REGION Network 34: Send preset command
   RUNG wire#powerrail
      Contact( #STC_tPH.x8 )
      wire#w1
      Contact( #STC_tMngSysReg.tST.xDone )
      wire#w2
      I_Contact( #STC_tMngSysReg.tST.xBusy )
      wire#w3
      I_Contact( #STC_tMngSysReg.tST.xError )
      S_Coil( #STC_tPH.x10 )
   END_RUNG
   RUNG wire#w1
      Contact( #STC_tMngSysReg.tST.xError )
   END_RUNG wire#w2
   RUNG wire#w3
      R_Coil( #STC_tPH.x8 )
   END_RUNG
   // the same network as SCL:
   #_w1 := #STC_tPH.x8 AND (#STC_tMngSysReg.tST.xDone OR #STC_tMngSysReg.tST.xError) AND NOT #STC_tMngSysReg.tST.xBusy;
   IF #_w1 AND NOT #STC_tMngSysReg.tST.xError THEN #STC_tPH.x10 := TRUE; END_IF;
   IF #_w1 THEN #STC_tPH.x8 := FALSE; END_IF;
END_REGION

REGION Network 35 (STL): Error during send ecoder value
         A     #STC_tMngSysReg.tST.xError;
         L     30;
         JC    Err;
END_REGION

REGION Network 36 (STL): Send preset command
         A     #STC_tPH.x10;
         JCN   PrE1;
         =     #STC_tMngSysReg.tST.xWrite_Request;

         L     #STC_tSYS_DATA.iPosPZD_MM;
         +     20;
         SLW   8;
         L     W#16#2;
         OW;
         T     #STC_tMngSysReg.tDATA.wRequest_refere_RequestID;
         L     #STC_tSYS_DATA.iPosPZD_MM;
         SLW   8;
         L     W#16#1;
         OW;
         T     #STC_tMngSysReg.tDATA.wAxis_NoOfParameters;
         L     W#16#1001;
         T     #STC_tMngSysReg.tDATA.wAttribute_NoOfElements;
         L     2507;
         T     #STC_tMngSysReg.tDATA.iParameter_number;
         L     W#16#0;
         T     #STC_tMngSysReg.tDATA.wSubindex;
         L     W#16#4201;
         T     #STC_tMngSysReg.tDATA.wFormat_NoOfValue;
         L     #STC_tSYS_DATA.iDiagAddress;
         T     #STC_tMngSysReg.tST.ID;
         L     47;
         T     #STC_tMngSysReg.tST.dINDEX;
         L     14;
         T     #STC_tMngSysReg.tST.uiLEN;

         L     DINT#2;
         SLD   16;
         T     #STC_tMngSysReg.tDATA.dwRegisterValue;

         CALL  #STC_tWriteRecord
         ( REQ    := #STC_tMngSysReg.tST.xWrite_Request,
           ID     := #STC_tMngSysReg.tST.ID,
           INDEX  := #STC_tMngSysReg.tST.dINDEX,
           LEN    := #STC_tMngSysReg.tST.uiLEN,
           DONE   := #STC_tMngSysReg.tST.xDone,
           BUSY   := #STC_tMngSysReg.tST.xBusy,
           ERROR  := #STC_tMngSysReg.tST.xError,
           STATUS := #STC_tMngSysReg.tST.dwSTATUS,
           RECORD := #STC_tMngSysReg.tDATA
         );
   PrE1: NOP   0;
END_REGION

REGION Network 37: Send saving preset command
   RUNG wire#powerrail
      Contact( #STC_tPH.x10 )
      wire#w1
      Contact( #STC_tMngSysReg.tST.xDone )
      wire#w2
      I_Contact( #STC_tMngSysReg.tST.xBusy )
      wire#w3
      I_Contact( #STC_tMngSysReg.tST.xError )
      S_Coil( #STC_tPH.x12 )
   END_RUNG
   RUNG wire#w1
      Contact( #STC_tMngSysReg.tST.xError )
   END_RUNG wire#w2
   RUNG wire#w3
      R_Coil( #STC_tPH.x10 )
   END_RUNG
   // the same network as SCL:
   #_w1 := #STC_tPH.x10 AND (#STC_tMngSysReg.tST.xDone OR #STC_tMngSysReg.tST.xError) AND NOT #STC_tMngSysReg.tST.xBusy;
   IF #_w1 AND NOT #STC_tMngSysReg.tST.xError THEN #STC_tPH.x12 := TRUE; END_IF;
   IF #_w1 THEN #STC_tPH.x10 := FALSE; END_IF;
END_REGION

REGION Network 38 (STL): Error during preset command
         A     #STC_tMngSysReg.tST.xError;
         L     31;
         JC    Err;
END_REGION

REGION Network 39 (STL): Send saving preset command
         A     #STC_tPH.x12;
         JCN   PrE2;
         =     #STC_tMngSysReg.tST.xWrite_Request;

         L     #STC_tSYS_DATA.iPosPZD_MM;
         +     30;
         SLW   8;
         L     W#16#2;
         OW;
         T     #STC_tMngSysReg.tDATA.wRequest_refere_RequestID;
         L     #STC_tSYS_DATA.iPosPZD_CU;
         SLW   8;
         L     W#16#1;
         OW;
         T     #STC_tMngSysReg.tDATA.wAxis_NoOfParameters;
         L     W#16#1001;
         T     #STC_tMngSysReg.tDATA.wAttribute_NoOfElements;
         L     977;
         T     #STC_tMngSysReg.tDATA.iParameter_number;
         L     W#16#0;
         T     #STC_tMngSysReg.tDATA.wSubindex;
         L     W#16#4201;
         T     #STC_tMngSysReg.tDATA.wFormat_NoOfValue;
         L     #STC_tSYS_DATA.iDiagAddress;
         T     #STC_tMngSysReg.tST.ID;
         L     47;
         T     #STC_tMngSysReg.tST.dINDEX;
         L     14;
         T     #STC_tMngSysReg.tST.uiLEN;

         L     DINT#1;
         SLD   16;
         T     #STC_tMngSysReg.tDATA.dwRegisterValue;

         CALL  #STC_tWriteRecord
         ( REQ    := #STC_tMngSysReg.tST.xWrite_Request,
           ID     := #STC_tMngSysReg.tST.ID,
           INDEX  := #STC_tMngSysReg.tST.dINDEX,
           LEN    := #STC_tMngSysReg.tST.uiLEN,
           DONE   := #STC_tMngSysReg.tST.xDone,
           BUSY   := #STC_tMngSysReg.tST.xBusy,
           ERROR  := #STC_tMngSysReg.tST.xError,
           STATUS := #STC_tMngSysReg.tST.dwSTATUS,
           RECORD := #STC_tMngSysReg.tDATA
         );
   PrE2: NOP   0;
END_REGION

REGION Network 40: End preset encoder
   RUNG wire#powerrail
      Contact( #STC_tPH.x12 )
      wire#w1
      Contact( #STC_tMngSysReg.tST.xDone )
      wire#w2
      I_Contact( #STC_tMngSysReg.tST.xBusy )
      wire#w3
      Coil( #STC_tPH.x14 )
   END_RUNG
   RUNG wire#w1
      Contact( #STC_tMngSysReg.tST.xError )
   END_RUNG wire#w2
   RUNG wire#w3
      R_Coil( #STC_tPH.x12 )
   END_RUNG
   // the same network as SCL:
   #STC_tPH.x14 := #STC_tPH.x12 AND (#STC_tMngSysReg.tST.xDone OR #STC_tMngSysReg.tST.xError) AND NOT #STC_tMngSysReg.tST.xBusy;
   IF #STC_tPH.x14 THEN #STC_tPH.x12 := FALSE; END_IF;
END_REGION

REGION Network 41 (STL): Error during saving preset command
         A     #STC_tMngSysReg.tST.xError;
         L     32;
         JC    Err;
END_REGION

REGION Network 42: Preset phases in progress
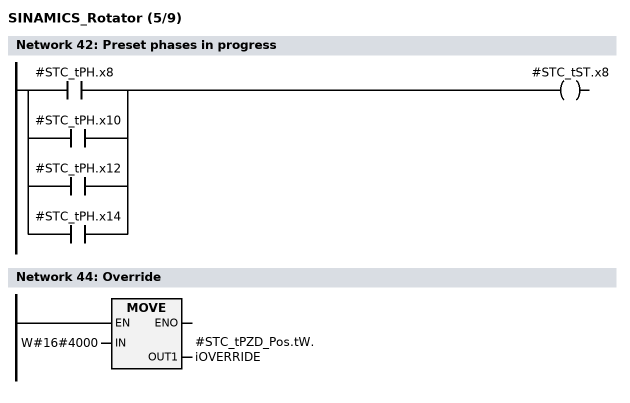
   RUNG wire#powerrail
      Contact( #STC_tPH.x8 )
      wire#w1
      Coil( #STC_tST.x8 )
   END_RUNG
   RUNG wire#powerrail
      Contact( #STC_tPH.x10 )
   END_RUNG wire#w1
   RUNG wire#powerrail
      Contact( #STC_tPH.x12 )
   END_RUNG wire#w1
   RUNG wire#powerrail
      Contact( #STC_tPH.x14 )
   END_RUNG wire#w1
   // the same network as SCL:
   #STC_tST.x8 := #STC_tPH.x8 OR #STC_tPH.x10 OR #STC_tPH.x12 OR #STC_tPH.x14;
END_REGION

REGION Network 43: #####_PARAMETERS_#####
END_REGION

REGION Network 44: Override
   RUNG wire#powerrail
      { S7_GenerateENO := "TRUE" } Move(in := W#16#4000, out1 => #STC_tPZD_Pos.tW.iOVERRIDE)
   END_RUNG
   // the same network as SCL:
   #STC_tPZD_Pos.tW.iOVERRIDE := W#16#4000;
END_REGION

REGION Network 45: Actual position filtered
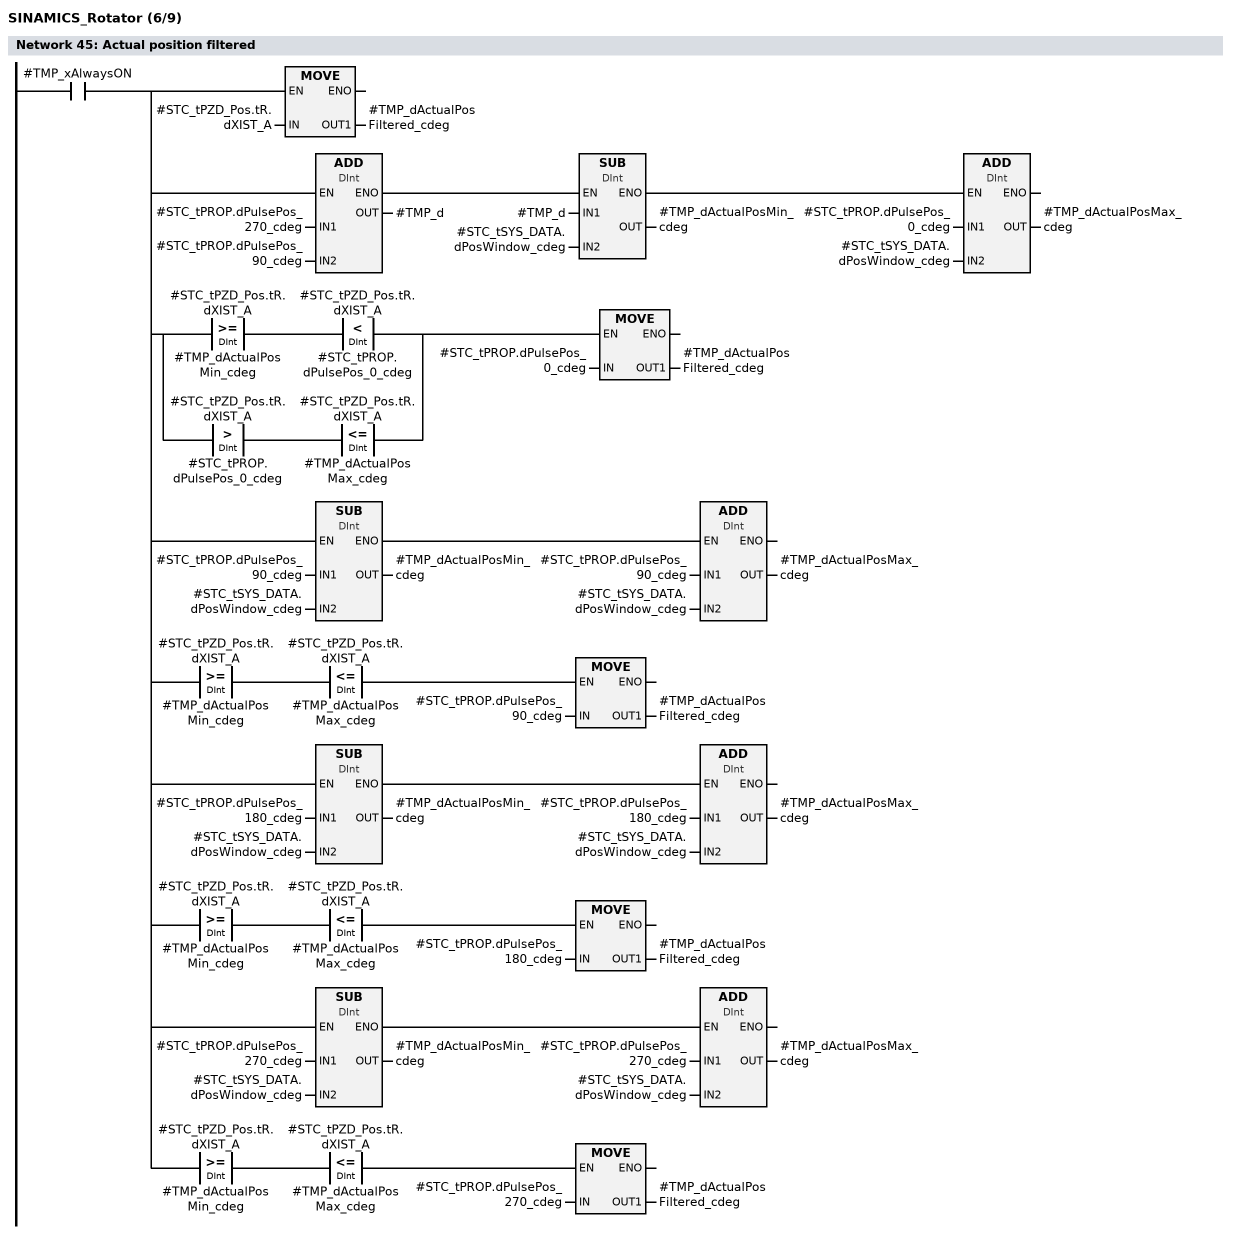
   RUNG wire#powerrail
      Contact( #TMP_xAlwaysON )
      wire#w1
      { S7_GenerateENO := "TRUE" } Move(in := #STC_tPZD_Pos.tR.dXIST_A, out1 => #TMP_dActualPosFiltered_cdeg)
   END_RUNG
   RUNG wire#w1
      { S7_Templates := "SrcType := DInt"; S7_GenerateENO := "TRUE" } Add(in1 := #STC_tPROP.dPulsePos_270_cdeg, in2 := #STC_tPROP.dPulsePos_90_cdeg, out => #TMP_d)
      { S7_Templates := "SrcType := DInt"; S7_GenerateENO := "TRUE" } Sub(in1 := #TMP_d, in2 := #STC_tSYS_DATA.dPosWindow_cdeg, out => #TMP_dActualPosMin_cdeg)
      { S7_Templates := "SrcType := DInt"; S7_GenerateENO := "TRUE" } Add(in1 := #STC_tPROP.dPulsePos_0_cdeg, in2 := #STC_tSYS_DATA.dPosWindow_cdeg, out => #TMP_dActualPosMax_cdeg)
   END_RUNG
   RUNG wire#w1
      { S7_Templates := "SrcType := DInt" } GE_Contact(in1 := #STC_tPZD_Pos.tR.dXIST_A, in2 := #TMP_dActualPosMin_cdeg)
      { S7_Templates := "SrcType := DInt" } LT_Contact(in1 := #STC_tPZD_Pos.tR.dXIST_A, in2 := #STC_tPROP.dPulsePos_0_cdeg)
      wire#w2
      { S7_GenerateENO := "TRUE" } Move(in := #STC_tPROP.dPulsePos_0_cdeg, out1 => #TMP_dActualPosFiltered_cdeg)
   END_RUNG
   RUNG wire#w1
      { S7_Templates := "SrcType := DInt" } GT_Contact(in1 := #STC_tPZD_Pos.tR.dXIST_A, in2 := #STC_tPROP.dPulsePos_0_cdeg)
      { S7_Templates := "SrcType := DInt" } LE_Contact(in1 := #STC_tPZD_Pos.tR.dXIST_A, in2 := #TMP_dActualPosMax_cdeg)
   END_RUNG wire#w2
   RUNG wire#w1
      { S7_Templates := "SrcType := DInt"; S7_GenerateENO := "TRUE" } Sub(in1 := #STC_tPROP.dPulsePos_90_cdeg, in2 := #STC_tSYS_DATA.dPosWindow_cdeg, out => #TMP_dActualPosMin_cdeg)
      { S7_Templates := "SrcType := DInt"; S7_GenerateENO := "TRUE" } Add(in1 := #STC_tPROP.dPulsePos_90_cdeg, in2 := #STC_tSYS_DATA.dPosWindow_cdeg, out => #TMP_dActualPosMax_cdeg)
   END_RUNG
   RUNG wire#w1
      { S7_Templates := "SrcType := DInt" } GE_Contact(in1 := #STC_tPZD_Pos.tR.dXIST_A, in2 := #TMP_dActualPosMin_cdeg)
      { S7_Templates := "SrcType := DInt" } LE_Contact(in1 := #STC_tPZD_Pos.tR.dXIST_A, in2 := #TMP_dActualPosMax_cdeg)
      { S7_GenerateENO := "TRUE" } Move(in := #STC_tPROP.dPulsePos_90_cdeg, out1 => #TMP_dActualPosFiltered_cdeg)
   END_RUNG
   RUNG wire#w1
      { S7_Templates := "SrcType := DInt"; S7_GenerateENO := "TRUE" } Sub(in1 := #STC_tPROP.dPulsePos_180_cdeg, in2 := #STC_tSYS_DATA.dPosWindow_cdeg, out => #TMP_dActualPosMin_cdeg)
      { S7_Templates := "SrcType := DInt"; S7_GenerateENO := "TRUE" } Add(in1 := #STC_tPROP.dPulsePos_180_cdeg, in2 := #STC_tSYS_DATA.dPosWindow_cdeg, out => #TMP_dActualPosMax_cdeg)
   END_RUNG
   RUNG wire#w1
      { S7_Templates := "SrcType := DInt" } GE_Contact(in1 := #STC_tPZD_Pos.tR.dXIST_A, in2 := #TMP_dActualPosMin_cdeg)
      { S7_Templates := "SrcType := DInt" } LE_Contact(in1 := #STC_tPZD_Pos.tR.dXIST_A, in2 := #TMP_dActualPosMax_cdeg)
      { S7_GenerateENO := "TRUE" } Move(in := #STC_tPROP.dPulsePos_180_cdeg, out1 => #TMP_dActualPosFiltered_cdeg)
   END_RUNG
   RUNG wire#w1
      { S7_Templates := "SrcType := DInt"; S7_GenerateENO := "TRUE" } Sub(in1 := #STC_tPROP.dPulsePos_270_cdeg, in2 := #STC_tSYS_DATA.dPosWindow_cdeg, out => #TMP_dActualPosMin_cdeg)
      { S7_Templates := "SrcType := DInt"; S7_GenerateENO := "TRUE" } Add(in1 := #STC_tPROP.dPulsePos_270_cdeg, in2 := #STC_tSYS_DATA.dPosWindow_cdeg, out => #TMP_dActualPosMax_cdeg)
   END_RUNG
   RUNG wire#w1
      { S7_Templates := "SrcType := DInt" } GE_Contact(in1 := #STC_tPZD_Pos.tR.dXIST_A, in2 := #TMP_dActualPosMin_cdeg)
      { S7_Templates := "SrcType := DInt" } LE_Contact(in1 := #STC_tPZD_Pos.tR.dXIST_A, in2 := #TMP_dActualPosMax_cdeg)
      { S7_GenerateENO := "TRUE" } Move(in := #STC_tPROP.dPulsePos_270_cdeg, out1 => #TMP_dActualPosFiltered_cdeg)
   END_RUNG
   // the same network as SCL:
   // ENO of a box is taken as its EN; it also drops when the box reports an error
   IF #TMP_xAlwaysON THEN
       #TMP_dActualPosFiltered_cdeg := #STC_tPZD_Pos.tR.dXIST_A;
       #TMP_d := #STC_tPROP.dPulsePos_270_cdeg + #STC_tPROP.dPulsePos_90_cdeg;
       #TMP_dActualPosMin_cdeg := #TMP_d - #STC_tSYS_DATA.dPosWindow_cdeg;
       #TMP_dActualPosMax_cdeg := #STC_tPROP.dPulsePos_0_cdeg + #STC_tSYS_DATA.dPosWindow_cdeg;
   END_IF;
   IF #TMP_xAlwaysON AND (((#STC_tPZD_Pos.tR.dXIST_A >= #TMP_dActualPosMin_cdeg) AND (#STC_tPZD_Pos.tR.dXIST_A < #STC_tPROP.dPulsePos_0_cdeg)) OR ((#STC_tPZD_Pos.tR.dXIST_A > #STC_tPROP.dPulsePos_0_cdeg) AND (#STC_tPZD_Pos.tR.dXIST_A <= #TMP_dActualPosMax_cdeg))) THEN
       #TMP_dActualPosFiltered_cdeg := #STC_tPROP.dPulsePos_0_cdeg;
   END_IF;
   IF #TMP_xAlwaysON THEN
       #TMP_dActualPosMin_cdeg := #STC_tPROP.dPulsePos_90_cdeg - #STC_tSYS_DATA.dPosWindow_cdeg;
       #TMP_dActualPosMax_cdeg := #STC_tPROP.dPulsePos_90_cdeg + #STC_tSYS_DATA.dPosWindow_cdeg;
   END_IF;
   IF #TMP_xAlwaysON AND (#STC_tPZD_Pos.tR.dXIST_A >= #TMP_dActualPosMin_cdeg) AND (#STC_tPZD_Pos.tR.dXIST_A <= #TMP_dActualPosMax_cdeg) THEN
       #TMP_dActualPosFiltered_cdeg := #STC_tPROP.dPulsePos_90_cdeg;
   END_IF;
   IF #TMP_xAlwaysON THEN
       #TMP_dActualPosMin_cdeg := #STC_tPROP.dPulsePos_180_cdeg - #STC_tSYS_DATA.dPosWindow_cdeg;
       #TMP_dActualPosMax_cdeg := #STC_tPROP.dPulsePos_180_cdeg + #STC_tSYS_DATA.dPosWindow_cdeg;
   END_IF;
   IF #TMP_xAlwaysON AND (#STC_tPZD_Pos.tR.dXIST_A >= #TMP_dActualPosMin_cdeg) AND (#STC_tPZD_Pos.tR.dXIST_A <= #TMP_dActualPosMax_cdeg) THEN
       #TMP_dActualPosFiltered_cdeg := #STC_tPROP.dPulsePos_180_cdeg;
   END_IF;
   IF #TMP_xAlwaysON THEN
       #TMP_dActualPosMin_cdeg := #STC_tPROP.dPulsePos_270_cdeg - #STC_tSYS_DATA.dPosWindow_cdeg;
       #TMP_dActualPosMax_cdeg := #STC_tPROP.dPulsePos_270_cdeg + #STC_tSYS_DATA.dPosWindow_cdeg;
   END_IF;
   IF #TMP_xAlwaysON AND (#STC_tPZD_Pos.tR.dXIST_A >= #TMP_dActualPosMin_cdeg) AND (#STC_tPZD_Pos.tR.dXIST_A <= #TMP_dActualPosMax_cdeg) THEN
       #TMP_dActualPosFiltered_cdeg := #STC_tPROP.dPulsePos_270_cdeg;
   END_IF;
END_REGION

REGION Network 46: Target selection
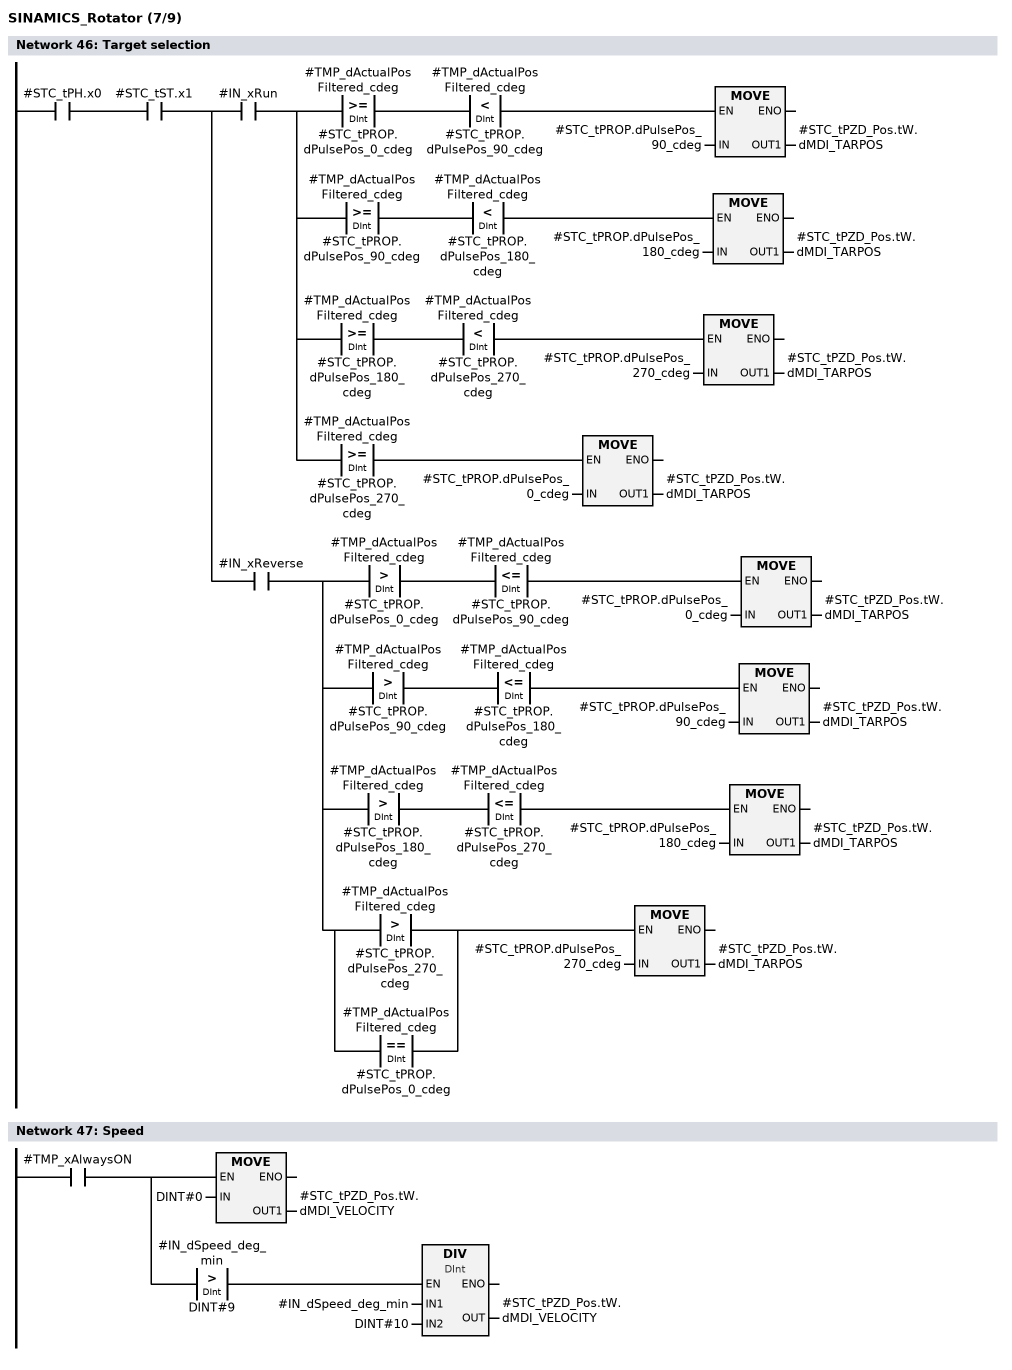
   RUNG wire#powerrail
      Contact( #STC_tPH.x0 )
      Contact( #STC_tST.x1 )
      wire#w1
      Contact( #IN_xRun )
      wire#w2
      { S7_Templates := "SrcType := DInt" } GE_Contact(in1 := #TMP_dActualPosFiltered_cdeg, in2 := #STC_tPROP.dPulsePos_0_cdeg)
      { S7_Templates := "SrcType := DInt" } LT_Contact(in1 := #TMP_dActualPosFiltered_cdeg, in2 := #STC_tPROP.dPulsePos_90_cdeg)
      { S7_GenerateENO := "TRUE" } Move(in := #STC_tPROP.dPulsePos_90_cdeg, out1 => #STC_tPZD_Pos.tW.dMDI_TARPOS)
   END_RUNG
   RUNG wire#w2
      { S7_Templates := "SrcType := DInt" } GE_Contact(in1 := #TMP_dActualPosFiltered_cdeg, in2 := #STC_tPROP.dPulsePos_90_cdeg)
      { S7_Templates := "SrcType := DInt" } LT_Contact(in1 := #TMP_dActualPosFiltered_cdeg, in2 := #STC_tPROP.dPulsePos_180_cdeg)
      { S7_GenerateENO := "TRUE" } Move(in := #STC_tPROP.dPulsePos_180_cdeg, out1 => #STC_tPZD_Pos.tW.dMDI_TARPOS)
   END_RUNG
   RUNG wire#w2
      { S7_Templates := "SrcType := DInt" } GE_Contact(in1 := #TMP_dActualPosFiltered_cdeg, in2 := #STC_tPROP.dPulsePos_180_cdeg)
      { S7_Templates := "SrcType := DInt" } LT_Contact(in1 := #TMP_dActualPosFiltered_cdeg, in2 := #STC_tPROP.dPulsePos_270_cdeg)
      { S7_GenerateENO := "TRUE" } Move(in := #STC_tPROP.dPulsePos_270_cdeg, out1 => #STC_tPZD_Pos.tW.dMDI_TARPOS)
   END_RUNG
   RUNG wire#w2
      { S7_Templates := "SrcType := DInt" } GE_Contact(in1 := #TMP_dActualPosFiltered_cdeg, in2 := #STC_tPROP.dPulsePos_270_cdeg)
      { S7_GenerateENO := "TRUE" } Move(in := #STC_tPROP.dPulsePos_0_cdeg, out1 => #STC_tPZD_Pos.tW.dMDI_TARPOS)
   END_RUNG
   RUNG wire#w1
      Contact( #IN_xReverse )
      wire#w3
      { S7_Templates := "SrcType := DInt" } GT_Contact(in1 := #TMP_dActualPosFiltered_cdeg, in2 := #STC_tPROP.dPulsePos_0_cdeg)
      { S7_Templates := "SrcType := DInt" } LE_Contact(in1 := #TMP_dActualPosFiltered_cdeg, in2 := #STC_tPROP.dPulsePos_90_cdeg)
      { S7_GenerateENO := "TRUE" } Move(in := #STC_tPROP.dPulsePos_0_cdeg, out1 => #STC_tPZD_Pos.tW.dMDI_TARPOS)
   END_RUNG
   RUNG wire#w3
      { S7_Templates := "SrcType := DInt" } GT_Contact(in1 := #TMP_dActualPosFiltered_cdeg, in2 := #STC_tPROP.dPulsePos_90_cdeg)
      { S7_Templates := "SrcType := DInt" } LE_Contact(in1 := #TMP_dActualPosFiltered_cdeg, in2 := #STC_tPROP.dPulsePos_180_cdeg)
      { S7_GenerateENO := "TRUE" } Move(in := #STC_tPROP.dPulsePos_90_cdeg, out1 => #STC_tPZD_Pos.tW.dMDI_TARPOS)
   END_RUNG
   RUNG wire#w3
      { S7_Templates := "SrcType := DInt" } GT_Contact(in1 := #TMP_dActualPosFiltered_cdeg, in2 := #STC_tPROP.dPulsePos_180_cdeg)
      { S7_Templates := "SrcType := DInt" } LE_Contact(in1 := #TMP_dActualPosFiltered_cdeg, in2 := #STC_tPROP.dPulsePos_270_cdeg)
      { S7_GenerateENO := "TRUE" } Move(in := #STC_tPROP.dPulsePos_180_cdeg, out1 => #STC_tPZD_Pos.tW.dMDI_TARPOS)
   END_RUNG
   RUNG wire#w3
      { S7_Templates := "SrcType := DInt" } GT_Contact(in1 := #TMP_dActualPosFiltered_cdeg, in2 := #STC_tPROP.dPulsePos_270_cdeg)
      wire#w4
      { S7_GenerateENO := "TRUE" } Move(in := #STC_tPROP.dPulsePos_270_cdeg, out1 => #STC_tPZD_Pos.tW.dMDI_TARPOS)
   END_RUNG
   RUNG wire#w3
      { S7_Templates := "SrcType := DInt" } EQ_Contact(in1 := #TMP_dActualPosFiltered_cdeg, in2 := #STC_tPROP.dPulsePos_0_cdeg)
   END_RUNG wire#w4
   // the same network as SCL:
   #_w1 := #STC_tPH.x0 AND #STC_tST.x1;
   #_w2 := #_w1 AND #IN_xRun;
   IF #_w2 AND (#TMP_dActualPosFiltered_cdeg >= #STC_tPROP.dPulsePos_0_cdeg) AND (#TMP_dActualPosFiltered_cdeg < #STC_tPROP.dPulsePos_90_cdeg) THEN
       #STC_tPZD_Pos.tW.dMDI_TARPOS := #STC_tPROP.dPulsePos_90_cdeg;
   END_IF;
   IF #_w2 AND (#TMP_dActualPosFiltered_cdeg >= #STC_tPROP.dPulsePos_90_cdeg) AND (#TMP_dActualPosFiltered_cdeg < #STC_tPROP.dPulsePos_180_cdeg) THEN
       #STC_tPZD_Pos.tW.dMDI_TARPOS := #STC_tPROP.dPulsePos_180_cdeg;
   END_IF;
   IF #_w2 AND (#TMP_dActualPosFiltered_cdeg >= #STC_tPROP.dPulsePos_180_cdeg) AND (#TMP_dActualPosFiltered_cdeg < #STC_tPROP.dPulsePos_270_cdeg) THEN
       #STC_tPZD_Pos.tW.dMDI_TARPOS := #STC_tPROP.dPulsePos_270_cdeg;
   END_IF;
   IF #_w2 AND (#TMP_dActualPosFiltered_cdeg >= #STC_tPROP.dPulsePos_270_cdeg) THEN
       #STC_tPZD_Pos.tW.dMDI_TARPOS := #STC_tPROP.dPulsePos_0_cdeg;
   END_IF;
   #_w3 := #_w1 AND #IN_xReverse;
   IF #_w3 AND (#TMP_dActualPosFiltered_cdeg > #STC_tPROP.dPulsePos_0_cdeg) AND (#TMP_dActualPosFiltered_cdeg <= #STC_tPROP.dPulsePos_90_cdeg) THEN
       #STC_tPZD_Pos.tW.dMDI_TARPOS := #STC_tPROP.dPulsePos_0_cdeg;
   END_IF;
   IF #_w3 AND (#TMP_dActualPosFiltered_cdeg > #STC_tPROP.dPulsePos_90_cdeg) AND (#TMP_dActualPosFiltered_cdeg <= #STC_tPROP.dPulsePos_180_cdeg) THEN
       #STC_tPZD_Pos.tW.dMDI_TARPOS := #STC_tPROP.dPulsePos_90_cdeg;
   END_IF;
   IF #_w3 AND (#TMP_dActualPosFiltered_cdeg > #STC_tPROP.dPulsePos_180_cdeg) AND (#TMP_dActualPosFiltered_cdeg <= #STC_tPROP.dPulsePos_270_cdeg) THEN
       #STC_tPZD_Pos.tW.dMDI_TARPOS := #STC_tPROP.dPulsePos_180_cdeg;
   END_IF;
   IF #_w3 AND ((#TMP_dActualPosFiltered_cdeg > #STC_tPROP.dPulsePos_270_cdeg) OR (#TMP_dActualPosFiltered_cdeg = #STC_tPROP.dPulsePos_0_cdeg)) THEN
       #STC_tPZD_Pos.tW.dMDI_TARPOS := #STC_tPROP.dPulsePos_270_cdeg;
   END_IF;
END_REGION

REGION Network 47: Speed
   RUNG wire#powerrail
      Contact( #TMP_xAlwaysON )
      wire#w1
      { S7_GenerateENO := "TRUE" } Move(in := DINT#0, out1 => #STC_tPZD_Pos.tW.dMDI_VELOCITY)
   END_RUNG
   RUNG wire#w1
      { S7_Templates := "SrcType := DInt" } GT_Contact(in1 := #IN_dSpeed_deg_min, in2 := DINT#9)
      { S7_Templates := "SrcType := DInt"; S7_GenerateENO := "TRUE" } Div(in1 := #IN_dSpeed_deg_min, in2 := DINT#10, out => #STC_tPZD_Pos.tW.dMDI_VELOCITY)
   END_RUNG
   // the same network as SCL:
   IF #TMP_xAlwaysON THEN #STC_tPZD_Pos.tW.dMDI_VELOCITY := DINT#0; END_IF;
   IF #TMP_xAlwaysON AND (#IN_dSpeed_deg_min > DINT#9) THEN
       #STC_tPZD_Pos.tW.dMDI_VELOCITY := #IN_dSpeed_deg_min / DINT#10;
   END_IF;
END_REGION

REGION Network 48: Acceleration
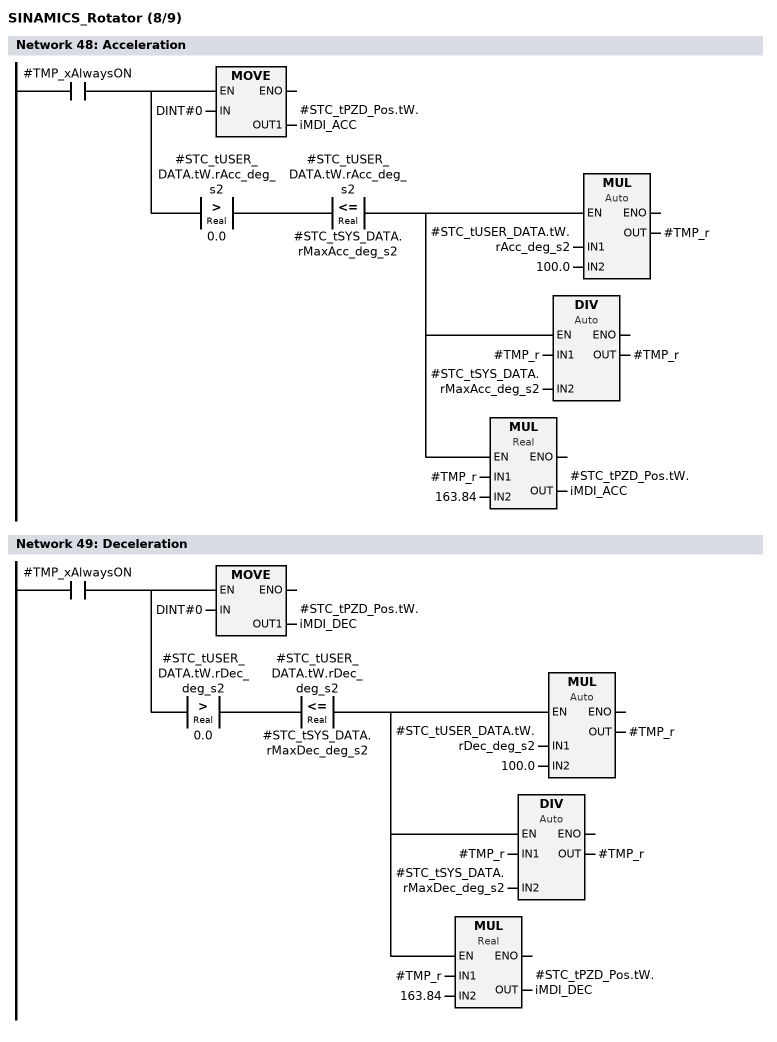
   RUNG wire#powerrail
      Contact( #TMP_xAlwaysON )
      wire#w1
      Move(in := DINT#0, out1 => #STC_tPZD_Pos.tW.iMDI_ACC)
   END_RUNG
   RUNG wire#w1
      { S7_Templates := "SrcType := Real" } GT_Contact(in1 := #STC_tUSER_DATA.tW.rAcc_deg_s2, in2 := 0.0)
      { S7_Templates := "SrcType := Real" } LE_Contact(in1 := #STC_tUSER_DATA.tW.rAcc_deg_s2, in2 := #STC_tSYS_DATA.rMaxAcc_deg_s2)
      wire#w2
      Mul(in1 := #STC_tUSER_DATA.tW.rAcc_deg_s2, in2 := 100.0, out => #TMP_r)
   END_RUNG
   RUNG wire#w2
      Div(in1 := #TMP_r, in2 := #STC_tSYS_DATA.rMaxAcc_deg_s2, out => #TMP_r)
   END_RUNG
   RUNG wire#w2
      { S7_Templates := "SrcType := Real" } Mul(in1 := #TMP_r, in2 := 163.84, out => #STC_tPZD_Pos.tW.iMDI_ACC)
   END_RUNG
   // the same network as SCL:
   IF #TMP_xAlwaysON THEN #STC_tPZD_Pos.tW.iMDI_ACC := DINT#0; END_IF;
   IF #TMP_xAlwaysON AND (#STC_tUSER_DATA.tW.rAcc_deg_s2 > 0.0) AND (#STC_tUSER_DATA.tW.rAcc_deg_s2 <= #STC_tSYS_DATA.rMaxAcc_deg_s2) THEN
       #TMP_r := #STC_tUSER_DATA.tW.rAcc_deg_s2 * 100.0;
       #TMP_r := #TMP_r / #STC_tSYS_DATA.rMaxAcc_deg_s2;
       #STC_tPZD_Pos.tW.iMDI_ACC := #TMP_r * 163.84;
   END_IF;
END_REGION

REGION Network 49: Deceleration
   RUNG wire#powerrail
      Contact( #TMP_xAlwaysON )
      wire#w1
      Move(in := DINT#0, out1 => #STC_tPZD_Pos.tW.iMDI_DEC)
   END_RUNG
   RUNG wire#w1
      { S7_Templates := "SrcType := Real" } GT_Contact(in1 := #STC_tUSER_DATA.tW.rDec_deg_s2, in2 := 0.0)
      { S7_Templates := "SrcType := Real" } LE_Contact(in1 := #STC_tUSER_DATA.tW.rDec_deg_s2, in2 := #STC_tSYS_DATA.rMaxDec_deg_s2)
      wire#w2
      Mul(in1 := #STC_tUSER_DATA.tW.rDec_deg_s2, in2 := 100.0, out => #TMP_r)
   END_RUNG
   RUNG wire#w2
      Div(in1 := #TMP_r, in2 := #STC_tSYS_DATA.rMaxDec_deg_s2, out => #TMP_r)
   END_RUNG
   RUNG wire#w2
      { S7_Templates := "SrcType := Real" } Mul(in1 := #TMP_r, in2 := 163.84, out => #STC_tPZD_Pos.tW.iMDI_DEC)
   END_RUNG
   // the same network as SCL:
   IF #TMP_xAlwaysON THEN #STC_tPZD_Pos.tW.iMDI_DEC := DINT#0; END_IF;
   IF #TMP_xAlwaysON AND (#STC_tUSER_DATA.tW.rDec_deg_s2 > 0.0) AND (#STC_tUSER_DATA.tW.rDec_deg_s2 <= #STC_tSYS_DATA.rMaxDec_deg_s2) THEN
       #TMP_r := #STC_tUSER_DATA.tW.rDec_deg_s2 * 100.0;
       #TMP_r := #TMP_r / #STC_tSYS_DATA.rMaxDec_deg_s2;
       #STC_tPZD_Pos.tW.iMDI_DEC := #TMP_r * 163.84;
   END_IF;
END_REGION

REGION Network 50: ################_MOTOR_MODULE_TELEGRAMS_ENDING_#################
END_REGION

REGION Network 51 (STL): Output copy motor module
   // Compute destination position
         L;
         LAR1;
   //byte 1 = 10h (FIXED for S7)
         L     B#16#10;
         T     B[AR1, P#0.0];
   //byte 2 = data type
         L     B#16#4;  //4 = word
         T     B[AR1, P#1.0];
   //byte 3 & 4 = number of element
         L     12;  //Production data
         T     W[AR1, P#2.0];
   //byte 5 & 6 = number of DB
         L     0;  //DB production data
         T     W[AR1, P#4.0];
   //byte 7 = memory area
         L     B#16#82;  //82h = Q (Output)
         T     B[AR1, P#6.0];
   //byte 8 & 9 = address. Bit 0,1,2 of tenth byte is bit offset
   //byte 7 = address (high). Valid value = 0-7. Bit 3,4,5,6,7 always 0
         L     #STC_tSYS_DATA.iIOAddress_MM;  //Item size
         SLW   3;
         T     W[AR1, P#8.0];
         SRD   16;
         AW    16#0007;
         T     B[AR1, P#7.0];

         CALL  BLKMOV
         ( SRCBLK  := #STC_tPZD_Pos.tW,
           RET_VAL := #TMP_iRetVal,
           DSTBLK  := #TMP_a
         );
END_REGION

REGION Network 52: #####_RETVAL_RESPONSE_#####
END_REGION

REGION Network 53 (STL): Initialize RetVal
         L     0;
         T     #OUT_iRetVal;
END_REGION

REGION Network 54: Warning messages
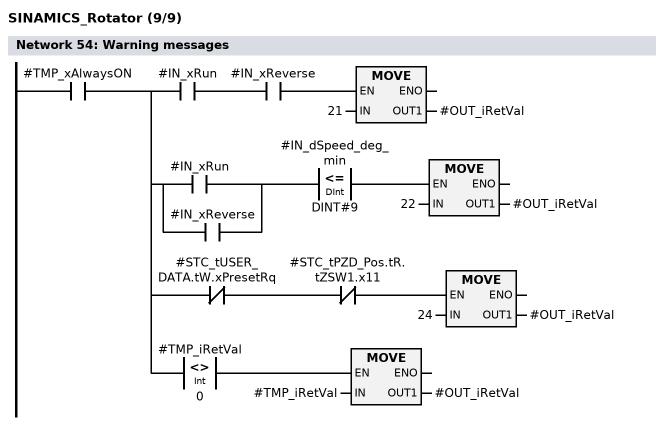
   RUNG wire#powerrail
      Contact( #TMP_xAlwaysON )
      wire#w1
      Contact( #IN_xRun )
      Contact( #IN_xReverse )
      { S7_GenerateENO := "TRUE" } Move(in := 21, out1 => #OUT_iRetVal)
   END_RUNG
   RUNG wire#w1
      Contact( #IN_xRun )
      wire#w2
      { S7_Templates := "SrcType := DInt" } LE_Contact(in1 := #IN_dSpeed_deg_min, in2 := DINT#9)
      { S7_GenerateENO := "TRUE" } Move(in := 22, out1 => #OUT_iRetVal)
   END_RUNG
   RUNG wire#w1
      Contact( #IN_xReverse )
   END_RUNG wire#w2
   RUNG wire#w1
      I_Contact( #STC_tUSER_DATA.tW.xPresetRq )
      I_Contact( #STC_tPZD_Pos.tR.tZSW1.x11 )
      { S7_GenerateENO := "TRUE" } Move(in := 24, out1 => #OUT_iRetVal)
   END_RUNG
   RUNG wire#w1
      { S7_Templates := "SrcType := Int" } NE_Contact(in1 := #TMP_iRetVal, in2 := 0)
      { S7_GenerateENO := "TRUE" } Move(in := #TMP_iRetVal, out1 => #OUT_iRetVal)
   END_RUNG
   // the same network as SCL:
   IF #TMP_xAlwaysON AND #IN_xRun AND #IN_xReverse THEN #OUT_iRetVal := 21; END_IF;
   IF #TMP_xAlwaysON AND (#IN_xRun OR #IN_xReverse) AND (#IN_dSpeed_deg_min <= DINT#9) THEN
       #OUT_iRetVal := 22;
   END_IF;
   IF #TMP_xAlwaysON AND NOT #STC_tUSER_DATA.tW.xPresetRq AND NOT #STC_tPZD_Pos.tR.tZSW1.x11 THEN
       #OUT_iRetVal := 24;
   END_IF;
   IF #TMP_xAlwaysON AND (#TMP_iRetVal <> 0) THEN #OUT_iRetVal := #TMP_iRetVal; END_IF;
END_REGION

REGION Network 55 (STL): Blocking messages
         JU    Rest;
   Err:  T     #OUT_iRetVal;
END_REGION

REGION Network 56 (STL): Reset input commands
   // R     #Run
   //       R     #Reverse
   //  
   // 
   //       L     L#0
   //       T     #Speed
   //       T     #USER_DATA.W.Acc
   //       T     #USER_DATA.W.Dec
   Rest: NOP   0;
   //    SET
   //    R     #IN_xDrive_EN
   //    R     #IN_xResetFaults
END_REGION

REGION Network 57 (STL): Restore AR1 & AR2 value
   //    L     #TMP_dOldValue_AR1
   //    LAR1
   //    L     #TMP_dOldValue_AR2
   //    LAR2
END_REGION
END_FUNCTION_BLOCK

